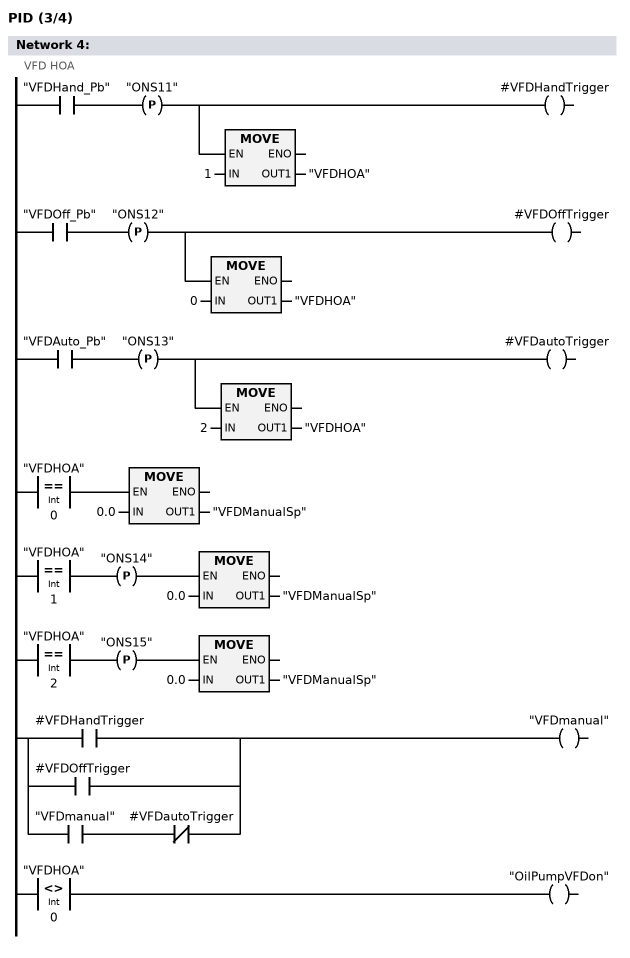
   RUNG wire#powerrail
      Contact( "VFDHand_Pb" )
      P_Trig( "ONS11" )
      wire#w1
      Coil( #VFDHandTrigger )
   END_RUNG
   RUNG wire#w1
      Move(in := 1, out1 => "VFDHOA")
   END_RUNG
   RUNG wire#powerrail
      Contact( "VFDOff_Pb" )
      P_Trig( "ONS12" )
      wire#w2
      Coil( #VFDOffTrigger )
   END_RUNG
   RUNG wire#w2
      Move(in := 0, out1 => "VFDHOA")
   END_RUNG
   RUNG wire#powerrail
      Contact( "VFDAuto_Pb" )
      P_Trig( "ONS13" )
      wire#w3
      Coil( #VFDautoTrigger )
   END_RUNG
   RUNG wire#w3
      Move(in := 2, out1 => "VFDHOA")
   END_RUNG
   RUNG wire#powerrail
      { S7_Templates := "SrcType := Int" } EQ_Contact(in1 := "VFDHOA", in2 := 0)
      Move(in := 0.0, out1 => "VFDManualSp")
   END_RUNG
   RUNG wire#powerrail
      { S7_Templates := "SrcType := Int" } EQ_Contact(in1 := "VFDHOA", in2 := 1)
      P_Trig( "ONS14" )
      Move(in := 0.0, out1 => "VFDManualSp")
   END_RUNG
   RUNG wire#powerrail
      { S7_Templates := "SrcType := Int" } EQ_Contact(in1 := "VFDHOA", in2 := 2)
      P_Trig( "ONS15" )
      Move(in := 0.0, out1 => "VFDManualSp")
   END_RUNG
   RUNG wire#powerrail
      Contact( #VFDHandTrigger )
      wire#w4
      Coil( "VFDmanual" )
   END_RUNG
   RUNG wire#powerrail
      Contact( #VFDOffTrigger )
   END_RUNG wire#w4
   RUNG wire#powerrail
      Contact( "VFDmanual" )
      I_Contact( #VFDautoTrigger )
   END_RUNG wire#w4
   RUNG wire#powerrail
      { S7_Templates := "SrcType := Int" } NE_Contact(in1 := "VFDHOA", in2 := 0)
      Coil( "OilPumpVFDon" )
   END_RUNG
   // the same network as SCL:
   #_w1 := "VFDHand_Pb" AND NOT "ONS11";   // rising edge
   "ONS11" := "VFDHand_Pb";
   #VFDHandTrigger := #_w1;
   IF #_w1 THEN "VFDHOA" := 1; END_IF;
   #_w2 := "VFDOff_Pb" AND NOT "ONS12";   // rising edge
   "ONS12" := "VFDOff_Pb";
   #VFDOffTrigger := #_w2;
   IF #_w2 THEN "VFDHOA" := 0; END_IF;
   #_w3 := "VFDAuto_Pb" AND NOT "ONS13";   // rising edge
   "ONS13" := "VFDAuto_Pb";
   #VFDautoTrigger := #_w3;
   IF #_w3 THEN "VFDHOA" := 2; END_IF;
   IF "VFDHOA" = 0 THEN "VFDManualSp" := 0.0; END_IF;
   #_w4 := "VFDHOA" = 1;
   #_w5 := #_w4 AND NOT "ONS14";   // rising edge
   "ONS14" := #_w4;
   IF #_w5 THEN "VFDManualSp" := 0.0; END_IF;
   #_w6 := "VFDHOA" = 2;
   #_w7 := #_w6 AND NOT "ONS15";   // rising edge
   "ONS15" := #_w6;
   IF #_w7 THEN "VFDManualSp" := 0.0; END_IF;
   "VFDmanual" := #VFDHandTrigger OR #VFDOffTrigger OR ("VFDmanual" AND NOT #VFDautoTrigger);
   "OilPumpVFDon" := "VFDHOA" <> 0;
END_REGION

REGION Network 5
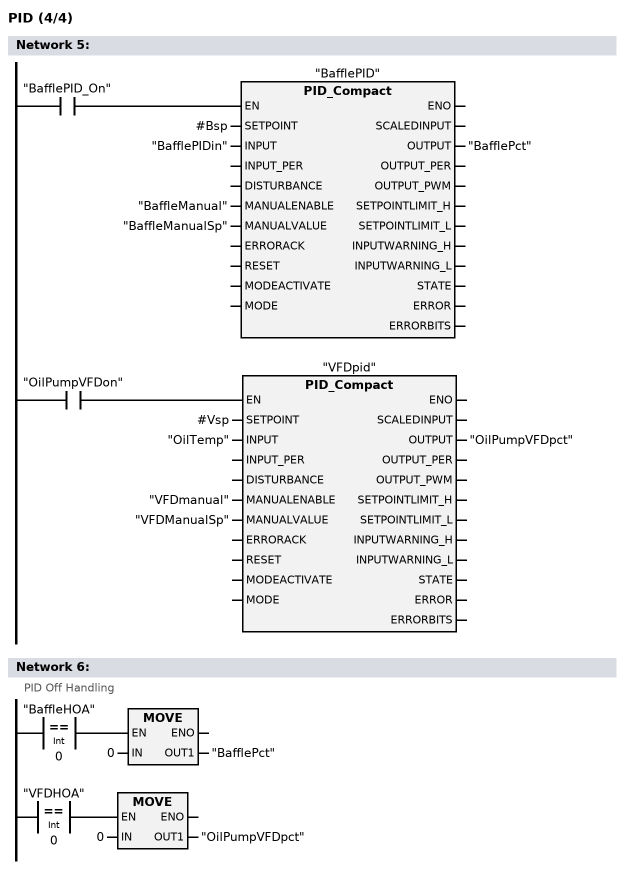
   IF "BafflePID_On" THEN
       "BafflePID"(Setpoint := #Bsp,   // PID_Compact
                   Input := "BafflePIDin",
                   ManualEnable := "BaffleManual",
                   ManualValue := "BaffleManualSp",
                   Output => "BafflePct");
   END_IF;
   IF "OilPumpVFDon" THEN
       "VFDpid"(Setpoint := #Vsp,   // PID_Compact
                Input := "OilTemp",
                ManualEnable := "VFDmanual",
                ManualValue := "VFDManualSp",
                Output => "OilPumpVFDpct");
   END_IF;
END_REGION

REGION Network 6
   // PID Off Handling
   RUNG wire#powerrail
      { S7_Templates := "SrcType := Int" } EQ_Contact(in1 := "BaffleHOA", in2 := 0)
      Move(in := 0, out1 => "BafflePct")
   END_RUNG
   RUNG wire#powerrail
      { S7_Templates := "SrcType := Int" } EQ_Contact(in1 := "VFDHOA", in2 := 0)
      Move(in := 0, out1 => "OilPumpVFDpct")
   END_RUNG
   // the same network as SCL:
   IF "BaffleHOA" = 0 THEN "BafflePct" := 0; END_IF;
   IF "VFDHOA" = 0 THEN "OilPumpVFDpct" := 0; END_IF;
END_REGION
END_ORGANIZATION_BLOCK

(* ===== HMI "HMI_RT_1" =====
system functions are stored by id; their names below are inferred from use
connection "1500PLC": S71200_TCP_IP, SCADA_S7_1500_OMS

HMI tags "Default tag table"
   "SystemStartPb" : Bool = PLC SystemStart_Pb AT %M65.2, 500 ms
   "SystemStopPb" : Bool = PLC SystemStop_Pb AT %M65.4, 500 ms
   "EStopAlarm" : Bool = PLC EStopAlarm AT %M49.3, 500 ms
   "BrakeFailureAlarm" : Bool = PLC BrakeFailureAlarm AT %M49.0, 500 ms
   "OverspeedAlarm" : Bool = PLC OverspeedAlarm AT %M48.4, 500 ms
   "OvercurrentAlarm" : Bool = PLC OvercurrentAlarm AT %M48.0, 500 ms
   "HighOilTempAlarm" : Bool = PLC HighOilTempAlarm AT %M48.2, 500 ms
   "HighOilFlowAlarm" : Bool = PLC OilHighFlowAlarm AT %M48.6, 500 ms
   "LowOilFlowAlarm" : Bool = PLC OilLowFlowAlarm AT %M5.6, 500 ms
   "AlarmSilence" : Bool = PLC AlarmSilence AT %M5.5, 500 ms
   "AlarmReset" : Bool = PLC AlarmReset AT %M5.4, 500 ms
   "BrakeEn" : Bool = PLC Brake_Out AT %M4.0, 500 ms
   "StationintlkEn" : Bool = PLC StationInterlock_Out AT %M3.1, 500 ms
   "VFDen" : Bool = PLC OilPumpVFDen_Out AT %M4.1, 500 ms
   "BaffleEn" : Int = PLC Baffle_Out AT %MW18, 500 ms
   "AlarmHornEn" : Bool = PLC AlarmHorn_Out AT %M3.0, 500 ms
   "BrakeHandPb" : Bool = PLC BrakeHand_Pb AT %M3.6, 500 ms
   "BrakeOffPb" : Bool = PLC BrakeOff_Pb AT %M3.5, 500 ms
   "BrakeAutoPb" : Bool = PLC BrakeAuto_Pb AT %M3.7, 500 ms
   "StationintlkHandPb" : Bool = PLC StationIntHand_Pb AT %M4.6, 500 ms
   "StationintlkOffPb" : Bool = PLC StationIntOff_Pb AT %M4.5, 500 ms
   "StationintlkAutoPb" : Bool = PLC StationIntAuto_Pb AT %M4.7, 500 ms
   "VFDhandPb" : Bool = PLC VFDHand_Pb AT %M99.3, 500 ms
   "VFDoffPb" : Bool = PLC VFDOff_Pb AT %M99.4, 500 ms
   "VFDautoPb" : Bool = PLC VFDAuto_Pb AT %M99.5, 500 ms
   "BaffleHandPb" : Bool = PLC BaffleHand_Pb AT %M98.5, 500 ms
   "BaffleOffPb" : Bool = PLC BaffleOff_Pb AT %M98.6, 500 ms
   "BaffleAutoPb" : Bool = PLC BaffleAuto_Pb AT %M98.4, 500 ms
   "AlarmHornHandPb" : Bool = PLC AlarmHornHand_Pb AT %M4.3, 500 ms
   "AlarmHornOffPb" : Bool = PLC AlarmHornOff_Pb AT %M4.2, 500 ms
   "AlarmHornAutoPb" : Bool = PLC AlarmHornAuto_Pb AT %M4.4, 500 ms
   "ModeInt" : Int = PLC ModeInt AT %MW118, 500 ms
   "BrakeHOA" : Int = PLC BrakeHoa AT %MW34, 500 ms
   "StationintlkHOA" : Int = PLC StationIntHoa AT %MW38, 500 ms
   "VFDhoa" : Int = PLC VFDHOA AT %MW108, 500 ms
   "BaffleHOA" : Int = PLC BaffleHOA AT %MW74, 500 ms
   "AlarmHornHOA" : Int = PLC AlarmHornHoa AT %MW36, 500 ms
   "HM_Minutes" : Int = PLC HM_Minutes AT %MW32, 500 ms
   "HM_Hours" : Int = PLC HM_Hours AT %MW114, 500 ms
   "HM_Days" : Int = PLC HM_Days AT %MW116, 500 ms
   "HM_ResetPb" : Bool = PLC ResetHourmeter_Pb AT %M106.7, 500 ms
   "FaultMode" : Bool = PLC FaultMode AT %M64.6, 500 ms
   "BrakeFailureDelay" : Int = PLC BrakeFailureDelay_Sp AT %MW62, 500 ms
   "OverCurrentSp" : Int = PLC OvercurrentSp AT %MW46, 500 ms
   "OvercurrentDelay" : Int = PLC OvercurrentDelay_Sp AT %MW44, 500 ms
   "OverspeedSp" : Int = PLC OverspeedSp AT %MW56, 500 ms
   "OverspeedDelay" : Int = PLC OverspeedDelay_Sp AT %MW54, 500 ms
   "HighOilTempSp" : Int = PLC HighOilTempSp AT %MW52, 500 ms
   "HighOilTempDelay" : Int = PLC HighOilTempDelay_Sp AT %MW50, 500 ms
   "HighOilFlowSp" : Int = PLC OilHHflowSp AT %MW60, 500 ms
   "HighOilFlowDelay" : Int = PLC OilHighFlowDelay_Sp AT %MW58, 500 ms
   "LowOilFlowSp" : Int = PLC OilLLflowSp AT %MW42, 500 ms
   "LowOilFlowDelay" : Int = PLC OilLowFlowDelay_Sp AT %MW40, 500 ms
   "WarmupOilTemp" : Int = PLC WarmupOilTemp AT %MW80, 500 ms
   "WarmUpDelay" : Int = PLC WarmupOilTempDelaySp AT %MW82, 500 ms
   "CurrentSp" : Int = PLC StabilizekWSp AT %MW86, 500 ms
   "StabilizeDelay" : Int = PLC StabilizeDelaySp AT %MW88, 500 ms
   "CooldownOilTemp" : Int = PLC CooldownOilTempSp AT %MW96, 500 ms
   "CooldownDelay" : Int = PLC CooldownDelaySp AT %MW92, 500 ms
   "VFDmanualSp" : Real = PLC VFDManualSp AT %MD110, 500 ms
   "BaffleManualSp" : Real = PLC BaffleManualSp AT %MD102, 500 ms
   "ProgramLanguage" : Int = PLC ProgLang AT %MW0, 500 ms
   "LADpb" : Bool = PLC PB_LAD AT %M2.1, 500 ms
   "FBDpb" : Bool = PLC PB_FBD AT %M2.5, 500 ms
   "SCLpb" : Bool = PLC PB_SCL AT %M2.6, 500 ms
   "STLpb" : Bool = PLC PB_STL AT %M2.7, 500 ms
   "Current" : Int = PLC Current AT %MW28, 500 ms
   "OilTemp" : Int = PLC OilTemp AT %MW20, 500 ms
   "OilFlow" : Int = PLC OilFlow AT %MW22, 500 ms
   "BafflePct" : Int = PLC BafflePct AT %MW10, 500 ms
   "VFDpct" : Int = PLC OilPumpVFDpct AT %MW8, 500 ms
   "RPM" : Int = PLC RPM AT %MW26, 500 ms
   "EStopNotify" : Bool = PLC EStopNotify AT %M49.4, 500 ms
   "BrakFailureNotify" : Bool = PLC BrakeFailureNotify AT %M49.1, 500 ms
   "OverspeedNotify" : Bool = PLC OverspeedNotify AT %M48.5, 500 ms
   "OvercurrentNotify" : Bool = PLC OvercurrentNotify AT %M48.1, 500 ms
   "HiTempNotify" : Bool = PLC HighOilTempNotify AT %M48.3, 500 ms
   "LoFlowNotify" : Bool = PLC OilLowFlowNotify AT %M5.7, 500 ms
   "HiFlowNotify" : Bool = PLC OilHighFlowNotify AT %M48.7, 500 ms

discrete alarms
   1: 'Estop open', class Errors, trigger "EStopNotify" bit 0
   2: 'Brake failed', class Errors, trigger "BrakFailureNotify" bit 0
   3: 'Overcurrent', class Errors, trigger "OvercurrentNotify" bit 0
   4: 'Overspeed', class Errors, trigger "OverspeedNotify" bit 0
   5: 'Hi oil flow', class Errors, trigger "HiFlowNotify" bit 0
   6: 'Lo oil flow', class Errors, trigger "LoFlowNotify" bit 0
   7: 'Hi oil temp', class Errors, trigger "HiTempNotify" bit 0

screen "Status" 500x500
   TextField "Text field_17" at 190,223 size 81x30; Text 'OFFLINE'
      Visibility <- "StationintlkEn"
   Button "Button_1" at 13,455 size 80x30; TextOff 'Main'
      on Click: ActivateScreen("Status", 0)
   Button "Button_2" at 109,455 size 80x30; TextOff 'Overview'
      on Click: ActivateScreen("Overview", 0)
   Button "Button_3" at 205,455 size 80x30; TextOff 'Alarms'
      on Click: ActivateScreen("Alarms", 0)
   Button "Button_4" at 301,455 size 80x30; TextOff 'Config'
      on Click: ActivateScreen("Config", 0)
   TextField "Text field_3" at 8,8 size 127x24; Text 'System Status'
   TextField "Text field_4" at 349,50 size 134x38; Text 'Idle Mode'
      Visibility <- "ModeInt"
   TextField "Text field_5" at 287,50 size 196x38; Text 'Warmup Mode'
      Visibility <- "ModeInt"
   TextField "Text field_6" at 290,50 size 193x38; Text 'Stabilize Mode'
      Visibility <- "ModeInt"
   TextField "Text field_7" at 254,50 size 229x38; Text 'Generation Mode'
      Visibility <- "ModeInt"
   TextField "Text field_8" at 271,50 size 212x38; Text 'Cooldown Mode'
      Visibility <- "ModeInt"
   TextField "Text field_9" at 340,294 size 145x26; Text 'Ladder Diagram'
      Visibility <- "ProgramLanguage"
   RoundButton "Round button_1" at 352,329 size 48x48; Text 'LAD'
      on PressLeft: SetBit("LADpb")
      on ReleaseLeft: ResetBit("LADpb")
   RoundButton "Round button_2" at 404,329 size 48x48; Text 'FBD'
      on PressLeft: SetBit("FBDpb")
      on ReleaseLeft: ResetBit("FBDpb")
   RoundButton "Round button_3" at 336,381 size 48x48; Text 'SCL'
      on PressLeft: SetBit("SCLpb")
      on ReleaseLeft: ResetBit("SCLpb")
   RoundButton "Round button_4" at 388,381 size 48x48; Text 'STL'
      on PressLeft: SetBit("STLpb")
      on ReleaseLeft: ResetBit("STLpb")
   TextField "Text field_10" at 354,294 size 130x26; Text 'Function Block'
      Visibility <- "ProgramLanguage"
   TextField "Text field_11" at 321,294 size 164x26; Text 'Structured Control'
      Visibility <- "ProgramLanguage"
   TextField "Text field_12" at 353,294 size 132x26; Text 'Statement List'
      Visibility <- "ProgramLanguage"
   RoundButton "Round button_5" at 34,335 size 94x94; Text 'START'
      on PressLeft: SetBit("SystemStartPb")
      on ReleaseLeft: ResetBit("SystemStartPb")
   RoundButton "Round button_6" at 153,337 size 94x94; Text 'STOP'
      on PressLeft: SetBit("SystemStopPb")
      on ReleaseLeft: ResetBit("SystemStopPb")
   IOField "I/O field_1" at 190,136 size 80x55; FormatPattern s99999
      ProcessValue <- "Current"
   TextField "Text field_13" at 104,151 size 73x24; Text 'Current:'
   TextField "Text field_14" at 278,151 size 28x24; Text 'kW'
   TextField "Text field_15" at 90,226 size 85x24; Text 'Interlock:'
   TextField "Text field_16" at 185,223 size 93x30; Text 'ENGAGED'
      Visibility <- "StationintlkEn"
   Group "Group_1" at 445,447 size 48x48
   Group "Group" at 445,447 size 48x48
      Visibility <- "FaultMode"
   TextField "Text field_2" at 456,462 size 25x19; Text 'OK!'
   TextField "Text field_1" at 445,461 size 47x19; Text 'Alarm!'

screen "Overview" 500x500
   Button "Button_1" at 13,455 size 80x30; TextOff 'Main'
      on Click: ActivateScreen("Status", 0)
   Button "Button_2" at 109,455 size 80x30; TextOff 'Overview'
      on Click: ActivateScreen("Overview", 0)
   Button "Button_3" at 205,455 size 80x30; TextOff 'Alarms'
      on Click: ActivateScreen("Alarms", 0)
   Button "Button_4" at 301,455 size 80x30; TextOff 'Config'
      on Click: ActivateScreen("Config", 0)
   TextField "Text field_3" at 8,8 size 154x24; Text 'System Overview'
   Group "Group_1" at 445,447 size 48x48
   Group "Group" at 445,447 size 48x48
      Visibility <- "FaultMode"
   GraphicView "Graphic view_1" at -14,32 size 520x324; Picture "System2_1"
   IOField "I/O field_1" at 8,332 size 63x38; FormatPattern 99999999
      ProcessValue <- "BafflePct"
   TextField "Text field_4" at 13,370 size 60x19; Text 'Baffle %'
   IOField "I/O field_2" at 238,332 size 63x38; FormatPattern 99999999
      ProcessValue <- "RPM"
   TextField "Text field_5" at 251,370 size 31x19; Text 'RPM'
   IOField "I/O field_3" at 189,122 size 63x38; FormatPattern 99999999
      ProcessValue <- "VFDpct"
   TextField "Text field_6" at 178,160 size 87x19; Text 'Oil Pump %'
   Group "Group_2" at 251,64 size 148x32
      Visibility <- "StationintlkEn"
   Group "Group_3" at 251,64 size 148x32
      Visibility <- "StationintlkEn"
   Group "Group_4" at 343,334 size 148x32
      Visibility <- "BrakeEn"
   Group "Group_5" at 343,334 size 148x32
      Visibility <- "BrakeEn"
   Group "Group_6" at 20,47 size 48x48
      Visibility <- "EStopAlarm"
   Group "Group_7" at 68,47 size 48x48
      Visibility <- "BrakeFailureAlarm"
   Group "Group_8" at 116,47 size 48x48
      Visibility <- "HighOilTempAlarm"
   Group "Group_9" at 20,95 size 48x48
      Visibility <- "HighOilFlowAlarm"
   Group "Group_10" at 68,95 size 48x48
      Visibility <- "LowOilFlowAlarm"
   Group "Group_11" at 116,95 size 48x48
      Visibility <- "OvercurrentAlarm"
   Group "Group_12" at 20,45 size 147x102
      Visibility <- "FaultMode"
   TextField "Text field_18" at 131,406 size 134x38; Text 'Idle Mode'
      Visibility <- "ModeInt"
   TextField "Text field_19" at 69,406 size 196x38; Text 'Warmup Mode'
      Visibility <- "ModeInt"
   TextField "Text field_20" at 72,406 size 193x38; Text 'Stabilize Mode'
      Visibility <- "ModeInt"
   TextField "Text field_21" at 36,406 size 229x38; Text 'Generation Mode'
      Visibility <- "ModeInt"
   TextField "Text field_22" at 53,406 size 212x38; Text 'Cooldown Mode'
      Visibility <- "ModeInt"
   Button "Button_5" at 403,388 size 80x30; TextOff 'Exit App'
      on Click: StopRuntime(0)
   IOField "I/O field_4" at 123,334 size 63x38; FormatPattern 99999999
      ProcessValue <- "OilTemp"
   TextField "Text field_23" at 120,372 size 66x19; Text 'Oil Temp'
   IOField "I/O field_5" at 318,391 size 63x38; FormatPattern 99999999
      ProcessValue <- "Current"
   TextField "Text field_24" at 336,429 size 22x19; Text 'kW'
   TextField "Text field_2" at 456,462 size 25x19; Text 'OK!'
   TextField "Text field_1" at 445,461 size 47x19; Text 'Alarm!'
   TextField "Text field_8" at 363,340 size 106x19; Text 'Brake Released'
   TextField "Text field_7" at 360,339 size 109x19; Text 'Brake Engaged!'
   TextField "Text field_10" at 262,70 size 128x19; Text 'Interlock Engaged'
   TextField "Text field_9" at 279,69 size 91x19; Text 'No Interlock!'
   TextField "Text field_11" at 23,61 size 41x19; Text 'EStop'
   TextField "Text field_12" at 73,61 size 39x19; Text 'Brake'
   TextField "Text field_13" at 120,61 size 41x19; Text 'Temp'
   TextField "Text field_14" at 25,111 size 38x17; Text 'HiFlow'
   TextField "Text field_15" at 71,111 size 42x17; Text 'LoFlow'
   TextField "Text field_16" at 129,111 size 22x19; Text 'kW'
   TextField "Text field_17" at 48,81 size 97x24; Text 'No Alarms.'

screen "Alarms" 500x500
   Button "Button_1" at 13,455 size 80x30; TextOff 'Main'
      on Click: ActivateScreen("Status", 0)
   Button "Button_2" at 109,455 size 80x30; TextOff 'Overview'
      on Click: ActivateScreen("Overview", 0)
   Button "Button_3" at 205,455 size 80x30; TextOff 'Alarms'
      on Click: ActivateScreen("Alarms", 0)
   Button "Button_4" at 301,455 size 80x30; TextOff 'Config'
      on Click: ActivateScreen("Config", 0)
   TextField "Text field_3" at 8,8 size 174x24; Text 'Alarm Management'
   AlarmControl "Alarm view_1" at 15,44 size 472x254
   RoundButton "Round button_1" at 264,347 size 75x75; Text 'Silence'
      on PressLeft: SetBit("AlarmSilence")
      on ReleaseLeft: ResetBit("AlarmSilence")
   RoundButton "Round button_2" at 352,347 size 75x75; Text 'Reset'
      on PressLeft: SetBit("AlarmReset")
      on ReleaseLeft: ResetBit("AlarmReset")
   TextField "Text field_4" at 284,316 size 116x22; Text 'Alarm Controls'
   Group "Group_2" at 43,333 size 48x48
      Visibility <- "EStopAlarm"
   Group "Group_3" at 91,333 size 48x48
      Visibility <- "BrakeFailureAlarm"
   Group "Group_4" at 139,333 size 48x48
      Visibility <- "HighOilTempAlarm"
   Group "Group_5" at 43,381 size 48x48
      Visibility <- "HighOilFlowAlarm"
   Group "Group_6" at 91,381 size 48x48
      Visibility <- "LowOilFlowAlarm"
   Group "Group_7" at 139,381 size 48x48
      Visibility <- "OvercurrentAlarm"
   Group "Group_8" at 43,331 size 147x102
      Visibility <- "FaultMode"
   Group "Group_1" at 445,447 size 48x48
   Group "Group" at 445,447 size 48x48
      Visibility <- "FaultMode"
   TextField "Text field_5" at 46,347 size 41x19; Text 'EStop'
   TextField "Text field_6" at 96,347 size 39x19; Text 'Brake'
   TextField "Text field_7" at 143,347 size 41x19; Text 'Temp'
   TextField "Text field_8" at 48,397 size 38x17; Text 'HiFlow'
   TextField "Text field_9" at 94,397 size 42x17; Text 'LoFlow'
   TextField "Text field_10" at 152,397 size 22x19; Text 'kW'
   TextField "Text field_11" at 71,367 size 97x24; Text 'No Alarms.'
   TextField "Text field_2" at 456,462 size 25x19; Text 'OK!'
   TextField "Text field_1" at 445,461 size 47x19; Text 'Alarm!'

screen "Config" 500x500
   TextField "Text field_2" at 456,462 size 25x19; Text 'OK!'
   Group "Group_1" at 445,447 size 48x48
   Button "Button_1" at 13,455 size 80x30; TextOff 'Main'
      on Click: ActivateScreen("Status", 0)
   Button "Button_2" at 109,455 size 80x30; TextOff 'Overview'
      on Click: ActivateScreen("Overview", 0)
   Button "Button_3" at 205,455 size 80x30; TextOff 'Alarms'
      on Click: ActivateScreen("Alarms", 0)
   Button "Button_4" at 301,455 size 80x30; TextOff 'Config'
      on Click: ActivateScreen("Config", 0)
   Group "Group" at 445,447 size 48x48
      Visibility <- "FaultMode"
   TextField "Text field_3" at 8,8 size 125x24; Text 'Configuration'
   Group "Group_3" at 327,209 size 166x237
   Group "Group_5" at 11,404 size 289x40
   TextField "Text field_21" at 387,11 size 98x19; Text 'HOA Controls'
   TextField "Text field_22" at 342,35 size 38x17; Text 'Horn'
   TextField "Text field_23" at 336,59 size 39x17; Text 'Brake'
   TextField "Text field_24" at 317,81 size 58x17; Text 'Interlock'
   TextField "Text field_25" at 323,105 size 119x17; Text 'Baffle'
   TextField "Text field_26" at 320,156 size 90x17; Text 'Oil Pump VFD'
   Button "Button_5" at 376,34 size 24x20; TextOff 'H'
      on PressLeft: SetBit("AlarmHornHandPb")
      on ReleaseLeft: ResetBit("AlarmHornHandPb")
   Button "Button_6" at 403,34 size 24x20; TextOff 'O'
      on PressLeft: SetBit("AlarmHornOffPb")
      on ReleaseLeft: ResetBit("AlarmHornOffPb")
   Button "Button_7" at 430,34 size 24x20; TextOff 'A'
      on PressLeft: SetBit("AlarmHornAutoPb")
      on ReleaseLeft: ResetBit("AlarmHornAutoPb")
   Rectangle "Rectangle_4" at 460,34 size 25x20
      Visibility <- "AlarmHornHOA"
   Rectangle "Rectangle_5" at 460,34 size 25x20
      Visibility <- "AlarmHornHOA"
   Rectangle "Rectangle_6" at 460,34 size 25x20
      Visibility <- "AlarmHornHOA"
   Rectangle "Rectangle_7" at 460,57 size 25x20
      Visibility <- "BrakeHOA"
   Rectangle "Rectangle_8" at 460,57 size 25x20
      Visibility <- "BrakeHOA"
   Rectangle "Rectangle_9" at 461,57 size 25x20
      Visibility <- "BrakeHOA"
   Rectangle "Rectangle_10" at 460,80 size 25x20
      Visibility <- "StationintlkHOA"
   Rectangle "Rectangle_11" at 460,80 size 25x20
      Visibility <- "StationintlkHOA"
   Rectangle "Rectangle_12" at 461,80 size 25x20
      Visibility <- "StationintlkHOA"
   Rectangle "Rectangle_13" at 393,131 size 25x20
      Visibility <- "BaffleHOA"
   Rectangle "Rectangle_14" at 393,131 size 25x20
      Visibility <- "BaffleHOA"
   Rectangle "Rectangle_15" at 394,131 size 25x20
      Visibility <- "BaffleHOA"
   Rectangle "Rectangle_16" at 392,179 size 25x20
      Visibility <- "VFDhoa"
   Rectangle "Rectangle_17" at 392,179 size 25x20
      Visibility <- "VFDhoa"
   Rectangle "Rectangle_18" at 393,179 size 25x20
      Visibility <- "VFDhoa"
   Button "Button_8" at 376,57 size 24x20; TextOff 'H'
      on PressLeft: SetBit("BrakeHandPb")
      on ReleaseLeft: ResetBit("BrakeHandPb")
   Button "Button_9" at 403,57 size 24x20; TextOff 'O'
      on PressLeft: SetBit("BrakeOffPb")
      on ReleaseLeft: ResetBit("BrakeOffPb")
   Button "Button_10" at 430,57 size 24x20; TextOff 'A'
      on PressLeft: SetBit("BrakeAutoPb")
      on ReleaseLeft: ResetBit("BrakeAutoPb")
   Button "Button_11" at 376,80 size 24x20; TextOff 'H'
      on PressLeft: SetBit("StationintlkHandPb")
      on ReleaseLeft: ResetBit("StationintlkHandPb")
   Button "Button_12" at 403,80 size 24x20; TextOff 'O'
      on PressLeft: SetBit("StationintlkOffPb")
      on ReleaseLeft: ResetBit("StationintlkOffPb")
   Button "Button_13" at 430,80 size 24x20; TextOff 'A'
      on PressLeft: SetBit("StationintlkAutoPb")
      on ReleaseLeft: ResetBit("StationintlkAutoPb")
   Button "Button_14" at 312,131 size 24x20; TextOff 'H'
      on PressLeft: SetBit("BaffleHandPb")
      on ReleaseLeft: ResetBit("BaffleHandPb")
   Button "Button_15" at 339,131 size 24x20; TextOff 'O'
      on PressLeft: SetBit("BaffleOffPb")
      on ReleaseLeft: ResetBit("BaffleOffPb")
   Button "Button_16" at 366,131 size 24x20; TextOff 'A'
      on PressLeft: SetBit("BaffleAutoPb")
      on ReleaseLeft: ResetBit("BaffleAutoPb")
   Button "Button_17" at 312,179 size 24x20; TextOff 'H'
      on PressLeft: SetBit("VFDhandPb")
      on ReleaseLeft: ResetBit("VFDhandPb")
   Button "Button_18" at 339,179 size 24x20; TextOff 'O'
      on PressLeft: SetBit("VFDoffPb")
      on ReleaseLeft: ResetBit("VFDoffPb")
   Button "Button_19" at 366,179 size 24x20; TextOff 'A'
      on PressLeft: SetBit("VFDautoPb")
      on ReleaseLeft: ResetBit("VFDautoPb")
   IOField "I/O field_16" at 423,119 size 64x32; FormatPattern s999999999.999
      ProcessValue <- "BaffleManualSp"
   IOField "I/O field_17" at 423,167 size 64x32; FormatPattern s999999999.999
      ProcessValue <- "VFDmanualSp"
   TextField "Text field_27" at 432,107 size 53x17; Text 'Manual Sp'
   TextField "Text field_28" at 432,155 size 53x17; Text 'Manual Sp'
   Group "Group_2" at 8,34 size 186x365
   TextField "Text field_1" at 445,461 size 47x19; Text 'Alarm!'
   IOField "I/O field_1" at 436,240 size 49x26; FormatPattern s99999
      ProcessValue <- "WarmupOilTemp"
   TextField "Text field_4" at 374,213 size 104x19; Text 'Process Values'
   TextField "Text field_5" at 340,242 size 93x17; Text 'Warmup Temp'
   TextField "Text field_6" at 340,277 size 92x17; Text 'Warmup Delay'
   TextField "Text field_7" at 350,311 size 82x17; Text 'Current (kW)'
   TextField "Text field_8" at 342,344 size 97x17; Text 'Stabilize Delay'
   TextField "Text field_9" at 332,378 size 100x17; Text 'Cooldown Temp'
   TextField "Text field_10" at 333,412 size 99x17; Text 'Cooldown Delay'
   IOField "I/O field_2" at 436,274 size 49x26; FormatPattern s99999
      ProcessValue <- "WarmUpDelay"
   IOField "I/O field_3" at 436,308 size 49x26; FormatPattern s99999
      ProcessValue <- "CurrentSp"
   IOField "I/O field_4" at 436,342 size 49x26; FormatPattern s99999
      ProcessValue <- "StabilizeDelay"
   IOField "I/O field_5" at 436,376 size 49x26; FormatPattern s99999
      ProcessValue <- "CooldownOilTemp"
   IOField "I/O field_6" at 436,410 size 49x26; FormatPattern s99999
      ProcessValue <- "CooldownDelay"
   IOField "I/O field_7" at 136,65 size 49x26; FormatPattern s99999
      ProcessValue <- "BrakeFailureDelay"
   TextField "Text field_11" at 88,38 size 94x19; Text 'Alarm Values'
   TextField "Text field_12" at 13,68 size 123x17; Text 'Brake Failure Delay'
   TextField "Text field_13" at 34,99 size 101x17; Text 'Overspeed RPM'
   TextField "Text field_14" at 27,127 size 107x17; Text 'Overspeed Delay'
   TextField "Text field_15" at 14,156 size 119x17; Text 'Overtemp Degrees'
   TextField "Text field_16" at 30,185 size 105x17; Text 'Overtemp Delay'
   IOField "I/O field_8" at 136,95 size 49x26; FormatPattern s99999
      ProcessValue <- "OverspeedSp"
   IOField "I/O field_9" at 136,124 size 49x26; FormatPattern s99999
      ProcessValue <- "OverspeedDelay"
   IOField "I/O field_10" at 136,153 size 49x26; FormatPattern s99999
      ProcessValue <- "HighOilTempSp"
   IOField "I/O field_11" at 136,183 size 49x26; FormatPattern s99999
      ProcessValue <- "HighOilTempDelay"
   TextField "Text field_17" at 51,215 size 84x17; Text 'Lo Flow GPM'
   TextField "Text field_18" at 42,245 size 92x17; Text 'Lo Flow Delay'
   TextField "Text field_19" at 51,275 size 84x17; Text 'Hi Flow GPM'
   TextField "Text field_20" at 46,305 size 87x17; Text 'Hi Flow Delay'
   IOField "I/O field_12" at 136,211 size 49x26; FormatPattern s99999
      ProcessValue <- "LowOilFlowSp"
   IOField "I/O field_13" at 136,241 size 49x26; FormatPattern s99999
      ProcessValue <- "LowOilFlowDelay"
   IOField "I/O field_14" at 136,271 size 49x26; FormatPattern s99999
      ProcessValue <- "HighOilFlowSp"
   IOField "I/O field_15" at 136,301 size 49x26; FormatPattern s99999
      ProcessValue <- "HighOilFlowDelay"
   TextField "Text field_33" at 30,335 size 102x17; Text 'Overcurrent kW'
   TextField "Text field_34" at 16,364 size 120x17; Text 'Overcurrent Delay'
   IOField "I/O field_21" at 136,332 size 49x26; FormatPattern s99999
      ProcessValue <- "OverCurrentSp"
   IOField "I/O field_22" at 136,362 size 49x26; FormatPattern s99999
      ProcessValue <- "OvercurrentDelay"
   IOField "I/O field_18" at 83,404 size 49x26; FormatPattern s99999
      ProcessValue <- "HM_Days"
   TextField "Text field_29" at 11,406 size 75x17; Text 'Hourmeter'
   Button "Button_20" at 251,404 size 49x25; TextOff 'RESET'
      on PressLeft: SetBit("HM_ResetPb")
      on ReleaseLeft: ResetBit("HM_ResetPb")
   IOField "I/O field_19" at 137,404 size 49x26; FormatPattern s99999
      ProcessValue <- "HM_Hours"
   IOField "I/O field_20" at 191,404 size 49x26; FormatPattern s99999
      ProcessValue <- "HM_Minutes"
   TextField "Text field_30" at 93,427 size 43x17; Text 'Days'
   TextField "Text field_31" at 202,427 size 43x17; Text 'Mins'
   TextField "Text field_32" at 143,427 size 43x17; Text 'Hours'
*)